// TIA Portal project "g" (V14)

(* hardware
DEVICE "S7-1200 station_1"  S7-1200 Station
   slot 0: "Rack_0"  S7-1200 Rack  Rack  V1.0
   slot 1: "PLC_1_test_mb_og_utv"  CPU 1217C DC/DC/DC  6ES7 217-1AG40-0XB0  V4.2
   slot 2: "DI 16x24VDC_1"  6ES7 221-1BH32-0XB0  V2.0
   slot 3: "CB 1241 (RS485)"  CB 1241 (RS485)  6ES7 241-1CH30-1XB0  V1.0
DEVICE "S7-1200 station_6"  S7-1200 Station
   slot 0: "Rack_0"  S7-1200 Rack  Rack  V1.0
   slot 1: "slib"  CPU 1211C DC/DC/DC  6ES7 211-1AE40-0XB0  V4.2
   slot 3: "CB 1241 (RS485)"  CB 1241 (RS485)  6ES7 241-1CH30-1XB0  V1.0
DEVICE "HMI"  TP900 Comfort
   slot 0: "TP900 Comfort"  TP900 Comfort  6AV2 124-0JC01-0AX0  14.0.1.0
   slot 1: "HMI_RT_2"  TP900 Comfort  6AV2 124-0JC01-0AX0  14.0.1.0
   slot 5: "HMI_2.IE_CP_1"  PROFINET Interface  14.0.1.0
      slot 1: "PROFINET Interface_1"  PROFINET Interface
         slot 1: "Port_1"  Port
         slot 2: "Port_2"  Port
   slot 7: "HMI_2.MPI/DP_CP_1"  MPI/DP Interface  14.0.1.0
DEVICE "S7-1200 station_2"  S7-1200 Station
   slot 0: "Rack_0"  S7-1200 Rack  Rack  V1.0
   slot 1: "PLC_1"  CPU 1211C DC/DC/DC  6ES7 211-1AE40-0XB0  V4.2
   slot 3: "CB 1241 (RS485)"  CB 1241 (RS485)  6ES7 241-1CH30-1XB0  V1.0
*)

// ===== PLC "PLC_1_test_mb_og_utv"  CPU 1217C DC/DC/DC =====

VAR_GLOBAL   // PLC tag table "Default tag table"
   "my_special_tag_name" AT %IW0 : Int;
   "tt" AT %I0.0 : Bool;
END_VAR

TYPE "mb_station_block_udt"
   STRUCT
      conf : Struct   // Configuration
         disable : Bool;   // Skip all queries
         read_only : Bool;   // Skip all write queries. (fc 5,6,15,16)
         max_comm_error : USInt := 2;   // Repeating erros before communication_error flag is set
         exec_x_quries : USInt := 1;   // Number of queries to be exec. at each loop.
      END_STRUCT;
      out : Struct   // Outputs
         error : Bool;   // All errors, including communication errors
         error_comm : Bool;   // only communication errors
         finnish : Bool;   // qid is handed over to next device.
      END_STRUCT;
      log : Struct   // Logging for development and debugging.
         connected_time : DTL;   // The time the device was connected to the bus
         disconnected_time : DTL;   // The time, if a device was disconnected to the bus
         done_cnt : UDInt;   // Successfully queries counter for this device
         error_comm_cnt : UDInt;   // Communication erros cnt.
         error_exception_cnt : UDInt;   // Failed queries counter for this device
         error_status : Word;   // Status code from mb_master or mb_client
         error_data_addr : UDInt;   // d_addr for last failed querie; handy for troubleshooting
      END_STRUCT;
      z : Struct   // Internal states.
         header_qid : UInt;   // qid value at device header
         comm_err_cnt : USInt;   // Repeating communication errors
         exec_cnt : USInt;   // Numb. of exec. q. this loop
         offset_qid : UInt := 1;   // Device query id.
         err_hold : Bool;   // Help var for .out.error
      END_STRUCT;
   END_STRUCT;
END_TYPE

// folder: mb_test

DATA_BLOCK "test_mb_t1_DB"   // DB1
{ S7_Optimized_Access := 'TRUE' }
VERSION : 0.1
// stored: InstanceOfName test_mb_1
"test_mb_1"
BEGIN
END_DATA_BLOCK

// folder: (top level)

FUNCTION_BLOCK "_read little"   // FB1, SCL
{ S7_Optimized_Access := 'TRUE' }
VERSION : 0.1
   VAR_INPUT
      mb_addr : USInt;
   END_VAR
   VAR_IN_OUT
      mb_query : "mb_query";
   END_VAR
   VAR
      sb : "mb_station_block_udt";
      data1 : Real;
      data2 : Real;
      data3 : Real;
      dommy : Bool;
      err : Int;
      pos : DInt;
   END_VAR
BEGIN

   #mb_query(mb_addr := 123,
             mode := #mb_query.c.read.holding_reg,
             data_addr := 12345,
             data_ptr := #dommy);

   IF #mb_query.Done THEN

       // #pos := "mb_pos"(mb_query := #mb_query, addr := 12345);
       #pos := UDINT_TO_DINT(12354 - #mb_query.data_addr) * 2;

       #err := READ_LITTLE(src_array := #mb_query.z.buffer,
                           dest_Variable => #data1,
                           pos := #pos);
       #err := READ_LITTLE(src_array := #mb_query.z.buffer,
                           dest_Variable => #data2,
                           pos := #pos);
       #err := READ_LITTLE(src_array := #mb_query.z.buffer,
                           dest_Variable => #data3,
                           pos := #pos);
   END_IF;
END_FUNCTION_BLOCK

FUNCTION_BLOCK "ABcounterEncoder"   // FB2, SCL
{ S7_Optimized_Access := 'TRUE' }
VERSION : 0.1
   VAR_INPUT
      pulsA : Bool;
      pulsB : Bool;
      reverce : Bool;
      factor : Real := 1.0;
   END_VAR
   VAR_OUTPUT
      pos : Real;
      uncertainPos : Bool;
   END_VAR
   VAR
      old : Struct
         pulsA : Bool;
         pulsB : Bool;
      END_STRUCT;
      cnt : DInt;
      firstScan : Bool := true;
   END_VAR
BEGIN
   // Position encoder based on two pulses which are 90 degree
   // phase shifted. 

   // TIP: Use a HSC (High speed conter) instead of this function
   // block. Using a hardware HSC will use less CPU resources.

   IF #firstScan THEN
       #uncertainPos := true;
   END_IF;

   IF #pulsA <> #old.pulsA OR #pulsB <> #old.pulsB THEN
       #cnt += SEL(G := #reverce XOR (
                    #pulsA <> NOT #old.pulsA
                    OR #pulsB <> NOT #old.pulsB),
                    IN0 := -1, IN1 := 1);
   END_IF;

   #pos := DINT_TO_REAL(#cnt) * #factor;
   #old.pulsA := #pulsA; 
   #old.pulsB := #pulsB; 
   #firstScan := false;
END_FUNCTION_BLOCK

FUNCTION_BLOCK "ABcounterCorrection"   // FB4, SCL
{ S7_Optimized_Access := 'TRUE' }
VERSION : 0.1
   VAR_INPUT
      switch : Bool;
      cnt : DInt;
   END_VAR
   VAR_OUTPUT
      deviation : DInt;
   END_VAR
   VAR_IN_OUT
      AB : "ABcounterEncoder";
   END_VAR
   VAR
      rtrig : R_TRIG;
   END_VAR
BEGIN
   #rtrig(CLK := #switch);

   // Log the max deviation
   IF NOT #AB.uncertainPos THEN
       #deviation := MAX(IN1 := #deviation, IN2 := ABS(#AB.cnt - #cnt));
   END_IF;

   IF #rtrig.Q THEN
       #AB.cnt := #cnt;
       #AB.uncertainPos := false;
   END_IF;
END_FUNCTION_BLOCK

FUNCTION "mb_get" : Void   // FC6, SCL
{ S7_Optimized_Access := 'TRUE' }
VERSION : 0.1
   VAR_INPUT
      addr : UDInt;
   END_VAR
   VAR_IN_OUT
      data_ptr : Variant;
      mb_query : "mb_query";
   END_VAR
   VAR_TEMP
      pos : DInt;
      err : Int;
   END_VAR
BEGIN
   IF #mb_query.z.run.qid_cnt = #mb_query.z.run.qid
       AND  #mb_query.Done
   THEN
       #pos := UDINT_TO_USINT(#addr - #mb_query.data_addr) * 2;
       #err := Deserialize(SRC_ARRAY := #mb_query.z.buffer,
                           DEST_VARIABLE => #data_ptr,
                           POS := #pos);
   END_IF;
END_FUNCTION

FUNCTION "mb_read_little_endian" : Void   // FC8, SCL
{ S7_Optimized_Access := 'TRUE' }
VERSION : 0.1
   VAR_INPUT
      addr : UDInt;
      n : USInt;
   END_VAR
   VAR_IN_OUT
      mb_query : "mb_query";
   END_VAR
   VAR_TEMP
      bo : Int;
      tmp : Byte;
      c : Int;
   END_VAR
BEGIN
   (* Read little endian:

      The function should be placed before a read query, and may be used 
      muliple times.

      "mb_read_little_endian"(addr := 100, n := 1, mb_query := #mb_query);
      "mb_read_little_endian"(addr := 200, n := 3, mb_query := #mb_query);

      #mb_query(mb_addr := ___MB_ADDR___,
                mode := #mb_query.c.read.holding_reg,
                data_addr := ___DATA_ADDR___,
                data_ptr := ___DATA___ );
   *) 

   IF #mb_query.z.run.qid_cnt + 1 = #mb_query.z.run.qid
       AND #mb_query.stat.done
       AND NOT #mb_query.z.run.insert
       AND NOT #mb_query.z.run.write // Read query
       AND #mb_query.conf.buffer_handler
   THEN
       #bo := UDINT_TO_INT(#addr - #mb_query.z.q.data_addr) * 2;

       FOR #c := #bo TO #bo + #n * 4 BY 4 DO
           #tmp := #mb_query.z.buffer[#bo + 0];
           #mb_query.z.buffer[#bo + 0] := #mb_query.z.buffer[#bo + 3];
           #mb_query.z.buffer[#bo + 3] := #tmp;

           #tmp := #mb_query.z.buffer[#bo + 1];
           #mb_query.z.buffer[#bo + 1] := #mb_query.z.buffer[#bo + 2];
           #mb_query.z.buffer[#bo + 2] := #tmp;
       END_FOR;
   END_IF;
END_FUNCTION

FUNCTION "mb_extra" : Bool   // FC9, SCL
{ S7_Optimized_Access := 'TRUE' }
VERSION : 0.1
   VAR_IN_OUT
      sb : "mb_station_block_udt";
      mb_query : "mb_query";
   END_VAR
BEGIN
   (* Example

   "mb_station_block_footer"(sb := #sb, mb_query := #mb_query);

   IF "mb_extra"(sb := #sb, mb_query := #mb_query) THEN
       #mb_query(mode := #mb_query.c.write.holding_reg,
                 data_addr := 12345,
                 data_ptr := ___CONFIG_PARAM___);
   END_IF;
   *)

   #mb_extra :=
   #mb_query.z.sb.sid = #mb_query.z.sb.sid_cnt
   AND NOT #sb.out.error_comm;
   // AND NOT #mb_query.stat.busy;
END_FUNCTION

ORGANIZATION_BLOCK "Main"   // OB1, SCL, ProgramCycle
TITLE = "Main Program Sweep (Cycle)"
{ S7_Optimized_Access := 'TRUE' }
VERSION : 0.1
   VAR_INPUT
      Initial_Call : Bool;   // Initial call of this OB
      Remanence : Bool;   // =True, if remanent data are available
   END_VAR
BEGIN
END_ORGANIZATION_BLOCK

// folder: mb_test

FUNCTION_BLOCK "test_mb_master"   // FB13, SCL
{ S7_Optimized_Access := 'TRUE' }
VERSION : 0.1
   VAR_INPUT
      REQ : Bool;
      MB_ADDR : UInt;
      MODE : USInt;
      DATA_ADDR : UDInt;
      DATA_LEN : UInt;
   END_VAR
   VAR_OUTPUT
      BUSY : Bool;
      ERROR : Bool;
      DONE : Bool;
      STATUS : Word;
   END_VAR
   VAR_IN_OUT
      DATA_PTR : "mb_internal_b";
   END_VAR
   VAR
      test : "test_mb_common";
   END_VAR
BEGIN
   #test(REQ := #REQ,
         MB_ADDR := #MB_ADDR,
         MODE := #MODE,
         DATA_ADDR := #DATA_ADDR,
         DATA_LEN := #DATA_LEN,
         BUSY => #BUSY,
         ERROR => #ERROR,
         DONE => #DONE,
         STATUS => #STATUS);
END_FUNCTION_BLOCK

FUNCTION_BLOCK "test_mb_common"   // FB14, SCL
{ S7_Optimized_Access := 'TRUE' }
VERSION : 0.1
   VAR_INPUT
      REQ : Bool;
      MB_ADDR : UInt;
      MODE : USInt;
      DATA_ADDR : UDInt;
      DATA_LEN : UInt;
   END_VAR
   VAR_OUTPUT
      BUSY : Bool;
      ERROR : Bool;
      DONE : Bool;
      STATUS : Word;
   END_VAR
   VAR
      fakeBus : Struct
         q : Struct
            mb_addr : UInt;
            mode : USInt;
            data_addr : UDInt;
            data_len : UInt;
         END_STRUCT;
         res : Struct
            done : Bool;
            error : Bool;
         END_STRUCT;
      END_STRUCT;
      state : Int;
      reset : Bool;
      cnt : Int;
   END_VAR
BEGIN
   // Fake query testing block

   CASE #state OF
       0:  // Wait for req.
           IF #REQ THEN
               #BUSY := true;
               #state += 1;
           END_IF;
           #cnt := 0; // Init cnt.

       1:  // Simulate some waite time
           #cnt += 1;
           #state += BOOL_TO_INT(#cnt > 5);

       2:  // Insert q-param to fake bus.
           #fakeBus.q.mb_addr := #MB_ADDR;
           #fakeBus.q.mode := #MODE;
           #fakeBus.q.data_addr := #DATA_ADDR;
           #fakeBus.q.data_len := #DATA_LEN;
           #cnt += 1; // The test device will insert resualt until next scan.

       3:  // Done or Eroor
           #fakeBus.q.mb_addr := 0;
           #fakeBus.q.mode := 0;
           #fakeBus.q.data_addr := 0;
           #fakeBus.q.data_len := 0;

           #DONE := #fakeBus.res.done;
           #ERROR := #fakeBus.res.error;
           IF NOT #DONE AND NOT #ERROR THEN
               #ERROR := true;
               #STATUS := 16#80C8;
           END_IF;
           #BUSY := false;
           #state := 0;
   END_CASE;

   IF #reset THEN
       #state := 0;
       #ERROR := false;
       #DONE := false;
       #BUSY := false;
   END_IF;

   #fakeBus.res.done := false;
   #fakeBus.res.error := false;
END_FUNCTION_BLOCK

FUNCTION_BLOCK "test_mb_client"   // FB15, SCL
{ S7_Optimized_Access := 'TRUE' }
VERSION : 0.1
   VAR_INPUT
      REQ : Bool;
      DISCONNECT : Bool;
      MB_MODE : USInt;
      DATA_ADDR : UDInt;
      DATA_LEN : UInt;
   END_VAR
   VAR_OUTPUT
      DONE : Bool;
      BUSY : Bool;
      ERROR : Bool;
      STATUS : Word;
   END_VAR
   VAR_IN_OUT
      MB_DATA_PTR : Variant;
      CONNECT : Variant;
   END_VAR
   VAR
      MB_Unit_ID : USInt;
      Connected : Bool;
      _ : Bool;
      test : "test_mb_common";
      cnt : UInt;
   END_VAR
BEGIN
   IF #DISCONNECT THEN
       #cnt := 0;
       #test.reset := true;
       #Connected := false;
   ELSE
       IF #cnt < 10 THEN
           #cnt += 1;
           #BUSY := true;
       ELSE
           #Connected := true;
           #test.reset := false;

       END_IF;
   END_IF;

   #test(REQ := #REQ,
         MB_ADDR := #MB_Unit_ID,
         MODE := #MB_MODE,
         DATA_ADDR := #DATA_ADDR,
         DATA_LEN := #DATA_LEN,
         BUSY => #BUSY,
         ERROR => #ERROR,
         DONE => #DONE,
         STATUS => #STATUS);
END_FUNCTION_BLOCK

FUNCTION_BLOCK "test_mb_1"   // FB16, SCL
{ S7_Optimized_Access := 'TRUE' }
VERSION : 0.1
   VAR_INPUT
      start : Bool;
   END_VAR
   VAR_OUTPUT
      DONE : Bool;
      ERROR : Bool;
   END_VAR
   VAR
      state : Int;
      old_state : Int;
      cnt : UInt;
      mx : UInt;
      mb_query : "mb_query";
      mb_master_1200_ctrl : "mb_master_1200_ctrl";
      mb_master_1500_ctrl : "mb_master_1200_ctrl";
      mb_client_ctrl : "mb_client_ctrl";
      mb_test_sb : Array[1..5] of "test_mb_sb1";
      mb_test_sb_fake : Array[1..5] of "test_mb_sb1_fake_device";
   END_VAR
   VAR_TEMP
      c : Int;
      dommy : Word;
   END_VAR
BEGIN
   CASE #state OF
       0:  // Wait for start signal.
           #state += BOOL_TO_INT(#start);
           #DONE := false;
           #ERROR := false;

       1:  // mb_master-1200
           #mb_test_sb[1].write1.real_1 := 0;
           #mb_test_sb[1].write1.real_2 := 0;
           #mb_test_sb[4].write1.real_1 := 0;
           #mb_test_sb[4].write1.real_2 := 0;
           #state += 1;
       2:  
           #mb_master_1200_ctrl(hardware_id := 1,
                                baud := 9600,
                                timeout := T#0s, // Auto
                                mb_query := #mb_query);

           #mb_test_sb[1].write1.real_1 := 12.34;
           #mb_test_sb[1].write1.real_2 := 56.78;
           #mb_test_sb[1]<?Sub?>(MB_ADDR := 1, mb_query := #mb_query);
           #mb_test_sb[2]<?Sub?>(MB_ADDR := 1, mb_query := #mb_query);
           #mb_test_sb[3]<?Sub?>(MB_ADDR := 1, mb_query := #mb_query);

           // Create some noice ...
           FOR #c := 0 TO UINT_TO_INT( #cnt ) MOD 7 DO
               #mb_query(mb_addr := 200, data_ptr := #dommy);
           END_FOR;

           #mb_test_sb[4].write1.real_1 := 90.12;
           #mb_test_sb[4].write1.real_2 := 34.56;
           #mb_test_sb[4]<?Sub?>(MB_ADDR := 1, mb_query := #mb_query);
           #mb_test_sb[5]<?Sub?>(MB_ADDR := 1, mb_query := #mb_query);

           FOR #c := 1 TO 5 DO
               #mb_test_sb_fake[#c]<?Sub?>(MB_ADDR := INT_TO_USINT(#c),
                                    mb_query := #mb_query,
                                    mb_test := #mb_master_1200_ctrl.master.TEST,
                                    mb_buffer := #mb_master_1200_ctrl.buffer.buffer);
           END_FOR;

           #state += BOOL_TO_INT(#cnt > 10000
                                 AND #mb_test_sb[1].read1.real_1 <> 12.34
                                 AND #mb_test_sb[1].read1.real_2 <> 56.78
                                 AND #mb_test_sb[4].read1.real_1 <> 90.12
                                 AND #mb_test_sb[4].read1.real_2 <> 34.56 );

           IF #mb_test_sb[1].read1.real_1 <> 12.34 AND #mb_test_sb[1].read1.real_1 <> 0
               OR #mb_test_sb[1].read1.real_2 <> 56.78 AND #mb_test_sb[1].read1.real_2 <> 0

               OR #mb_test_sb[4].read1.real_1 <> 90.12 AND #mb_test_sb[4].read1.real_1 <> 0
               OR #mb_test_sb[4].read1.real_2 <> 34.56 AND #mb_test_sb[4].read1.real_2 <> 0
           THEN
               #state := -1; // Error
           END_IF;

       3:  // 1500
           #mb_test_sb[3].read1.real_1 := 0;
           #state += 1;
       4:
           #mb_master_1500_ctrl(hardware_id := 1,
                                baud := 9600,
                                timeout := T#300ms,
                                mb_query := #mb_query);

           #mb_test_sb[3].write1.real_1 := 98.76;

           FOR #c := 1 TO 5 DO
               #mb_test_sb[#c]<?Sub?>(MB_ADDR := INT_TO_USINT(#c),
                               mb_query := #mb_query);
           END_FOR;

           #mb_test_sb_fake[2]<?Sub?>(MB_ADDR := INT_TO_USINT(2),
                               mb_query := #mb_query,
                               mb_test := #mb_master_1500_ctrl.master.TEST,
                               mb_buffer := #mb_master_1500_ctrl.buffer.buffer);

           #state += BOOL_TO_INT(#cnt > 10000 AND #mb_test_sb[3].read1.real_1 <> 98.76 );

           IF #mb_test_sb[3].read1.real_1 <> 98.76 AND #mb_test_sb[3].read1.real_1 <> 0 THEN
               #state := -2; // Error
               #state += 1;
           END_IF;

       5:  // Client
           #mb_test_sb[2].read1.real_1 := 0;
       6:
           #mb_client_ctrl(mb_query := #mb_query);

           #mb_test_sb[2].write1.real_1 := 0.000076;

           FOR #c := 1 TO 5 DO
               #mb_test_sb[#c]<?Sub?>(MB_ADDR := INT_TO_USINT(#c), mb_query := #mb_query);
           END_FOR;

           #mb_test_sb_fake[2]<?Sub?>(MB_ADDR := INT_TO_USINT(2),
                               mb_query := #mb_query,
                               mb_test := #mb_master_1200_ctrl.master.TEST,
                               mb_buffer := #mb_master_1200_ctrl.buffer.buffer);

           #state += BOOL_TO_INT(#cnt > 10000
                                 AND #mb_test_sb[2].read1.real_1 <> 0.000076);

           IF #mb_test_sb[2].read1.real_1 <> 0.000076 AND #mb_test_sb[2].read1.real_1 <> 0 THEN
               #state := -2; // Error
           END_IF;

       7:
           #DONE := true;
   END_CASE;

   #cnt += 1;
   IF #old_state <> #state THEN
       #cnt := 0;
   END_IF;
   #old_state := #state;

   #ERROR := #state < 0;
END_FUNCTION_BLOCK

FUNCTION_BLOCK "test_mb_comm_load"   // FB17, SCL
{ S7_Optimized_Access := 'TRUE' }
VERSION : 0.1
   VAR_INPUT
      REQ : Bool;
      PORT : Port;
      BAUD : UInt;
      PARITY : UInt;
      RESP_TO : UInt;
   END_VAR
   VAR_OUTPUT
      DONE : Bool;
      ERROR : Bool;
   END_VAR
   VAR_IN_OUT
      MB_DB : Variant;
   END_VAR
   VAR
      MB_COMM_LOAD_Instance : MB_COMM_LOAD;
      "1500" : Bool;
   END_VAR
BEGIN

   IF #"1500" THEN
       #DONE := false;
   END_IF;

   IF #REQ  
       AND #PORT <> 0 AND #BAUD <> 0 AND #PARITY <> 0 AND #RESP_TO <> 0
   THEN
       #DONE := true;
   END_IF;

   #ERROR := NOT #DONE;
END_FUNCTION_BLOCK

FUNCTION_BLOCK "test_mb_sb1_fake_device"   // FB18, SCL
{ S7_Optimized_Access := 'TRUE' }
VERSION : 0.1
   VAR_INPUT
      MB_ADDR : UInt;
   END_VAR
   VAR_IN_OUT
      mb_query : "mb_query";
      mb_test : "test_mb_common";
      mb_buffer : Array[0..250] of Byte;
   END_VAR
   VAR
      fakeBus : Struct
         q : Struct
            mb_addr : UInt;
            mode : USInt;
            data_addr : UDInt;
            data_len : UInt;
         END_STRUCT;
         res : Struct
            done : Bool;
            error : Bool;
         END_STRUCT;
      END_STRUCT;
      read1 : Struct
         real_1 : Real;
         real_2 : Real;
         udint_1 : UDInt;
      END_STRUCT;
      read2 : Struct
         x00 : Bool;
         x01 : Bool;
         x02 : Bool;
         x03 : Bool;
         x04 : Bool;
         x05 : Bool;
         x06 : Bool;
         x07 : Bool;
         x08 : Bool;
         x09 : Bool;
         x10 : Bool;
         x11 : Bool;
         x12 : Bool;
         x13 : Bool;
         x14 : Bool;
         x15 : Bool;
      END_STRUCT;
      write1 : Struct
         real_2 : Real;
         udint_1 : UDInt;
         real_1 : Real;
      END_STRUCT;
      sb : "mb_station_block_udt";
   END_VAR
   VAR_TEMP
      pos : DInt;
      "e" : Int;
   END_VAR
BEGIN
   // Simulating a device 

   IF #mb_test.fakeBus.q.mb_addr = #MB_ADDR 
       AND #mb_test.fakeBus.q.data_len > 1
   THEN
       // Read 1
       IF #mb_test.fakeBus.q.mode = #mb_query.c.read.holding_reg
           AND #mb_test.fakeBus.q.data_addr = 123
       THEN
           #"e" := Serialize(SRC_VARIABLE := #read1, DEST_ARRAY => #mb_buffer, POS := #pos);
           #mb_test.fakeBus.res.done := #"e" = 0 AND #pos / 2 = #mb_test.fakeBus.q.data_len;
       END_IF;

       // Read 2
       IF #mb_test.fakeBus.q.mode = #mb_query.c.read.holding_reg
           AND #mb_test.fakeBus.q.data_addr = 456
       THEN
           #"e" := Serialize(SRC_VARIABLE := #read2, DEST_ARRAY => #mb_buffer, POS := #pos);
           #mb_test.fakeBus.res.done := #"e" = 0 AND #pos / 2 = #mb_test.fakeBus.q.data_len;
       END_IF;

       // Write 1
       IF #mb_test.fakeBus.q.mode = #mb_query.c.write.holding_reg
           AND #mb_test.fakeBus.q.data_addr = 789
       THEN
           #"e" := Deserialize(SRC_ARRAY := #mb_buffer, DEST_VARIABLE => #write1, POS := #pos);
           #mb_test.fakeBus.res.done := #"e" = 0 AND #pos / 2 = #mb_test.fakeBus.q.data_len;
       END_IF;
   END_IF;

   #mb_test.fakeBus.res.error := NOT #mb_test.fakeBus.res.done;

   #read1.real_1 := #write1.real_1;
   #read1.real_2 := #write1.real_2;
   #read1.udint_1 := #write1.udint_1;
END_FUNCTION_BLOCK

FUNCTION_BLOCK "test_mb_sb1"   // FB19, SCL
{ S7_Optimized_Access := 'TRUE' }
VERSION : 0.1
   VAR_INPUT
      MB_ADDR : UInt;
   END_VAR
   VAR_IN_OUT
      mb_query : "mb_query";
   END_VAR
   VAR
      fakeBus : Struct
         q : Struct
            mb_addr : UInt;
            mode : USInt;
            data_addr : UDInt;
            data_len : UInt;
         END_STRUCT;
         res : Struct
            done : Bool;
            error : Bool;
         END_STRUCT;
      END_STRUCT;
      read1 : Struct
         real_1 : Real;
         real_2 : Real;
         udint_1 : UDInt;
      END_STRUCT;
      read2 : Struct
         x00 : Bool;
         x01 : Bool;
         x02 : Bool;
         x03 : Bool;
         x04 : Bool;
         x05 : Bool;
         x06 : Bool;
         x07 : Bool;
         x08 : Bool;
         x09 : Bool;
         x10 : Bool;
         x11 : Bool;
         x12 : Bool;
         x13 : Bool;
         x14 : Bool;
         x15 : Bool;
      END_STRUCT;
      write1 : Struct
         real_2 : Real;
         udint_1 : UDInt;
         real_1 : Real;
      END_STRUCT;
      sb : "mb_station_block_udt";
      q1_done_cnt : UDInt;
      q2_done_cnt : UDInt;
      q3_done_cnt : UDInt;
   END_VAR
BEGIN
   // Testing device

   "mb_station_block_header"(sb := #sb, mb_query := #mb_query);
   #mb_query.mb_addr := #MB_ADDR;

   #mb_query(mode := #mb_query.c.read.holding_reg,
             data_addr := 123,
             data_ptr := #read1);
   #q1_done_cnt += BOOL_TO_UDINT(#mb_query.Done);

   #mb_query(mode := #mb_query.c.read.holding_reg,
             data_addr := 456,
             data_ptr := #read2);
   #q2_done_cnt += BOOL_TO_UDINT(#mb_query.Done);

   #mb_query(mode := #mb_query.c.write.holding_reg,
             data_addr := 789,
             data_ptr := #write1);
   #q3_done_cnt += BOOL_TO_UDINT(#mb_query.Done);

   "mb_station_block_footer"(sb := #sb, mb_query := #mb_query);
END_FUNCTION_BLOCK

FUNCTION_BLOCK "test_mb_sb2"   // FB20, SCL
{ S7_Optimized_Access := 'TRUE' }
VERSION : 0.1
   VAR_INPUT
      MB_ADDR : UInt;
   END_VAR
   VAR_IN_OUT
      mb_query : "mb_query";
   END_VAR
   VAR
      fakeBus : Struct
         q : Struct
            mb_addr : UInt;
            mode : USInt;
            data_addr : UDInt;
            data_len : UInt;
         END_STRUCT;
         res : Struct
            done : Bool;
            error : Bool;
         END_STRUCT;
      END_STRUCT;
      read1 : Struct
         real_1 : Real;
         real_2 : Real;
         udint_1 : UDInt;
      END_STRUCT;
      read2 : Struct
         x00 : Bool;
         x01 : Bool;
         x02 : Bool;
         x03 : Bool;
         x04 : Bool;
         x05 : Bool;
         x06 : Bool;
         x07 : Bool;
         x08 : Bool;
         x09 : Bool;
         x10 : Bool;
         x11 : Bool;
         x12 : Bool;
         x13 : Bool;
         x14 : Bool;
         x15 : Bool;
      END_STRUCT;
      write1 : Struct
         real_2 : Real;
         udint_1 : UDInt;
         real_1 : Real;
      END_STRUCT;
      sb : "mb_station_block_udt";
      q1_done_cnt : UDInt;
      q2_done_cnt : UDInt;
      q3_done_cnt : UDInt;
   END_VAR
BEGIN
   // Testing device

   "mb_station_block_header"(sb := #sb, mb_query := #mb_query);
   #mb_query.mb_addr := #MB_ADDR;

   #mb_query(mode := #mb_query.c.read.holding_reg,
             data_addr := 123,
             data_ptr := #read1);
   #q1_done_cnt += BOOL_TO_UDINT(#mb_query.Done);

   #mb_query(mode := #mb_query.c.read.holding_reg,
             data_addr := 456,
             data_ptr := #read2);
   #q2_done_cnt += BOOL_TO_UDINT(#mb_query.Done);

   #mb_query(mode := #mb_query.c.write.holding_reg,
             data_addr := 789,
             data_ptr := #write1);
   #q3_done_cnt += BOOL_TO_UDINT(#mb_query.Done);

   "mb_station_block_footer"(sb := #sb, mb_query := #mb_query);
END_FUNCTION_BLOCK

FUNCTION_BLOCK "test_mb_sb2_fake_device"   // FB21, SCL
{ S7_Optimized_Access := 'TRUE' }
VERSION : 0.1
   VAR_INPUT
      MB_ADDR : UInt;
   END_VAR
   VAR_IN_OUT
      mb_query : "mb_query";
      mb_test : "test_mb_common";
      mb_buffer : Array[0..250] of Byte;
   END_VAR
   VAR
      fakeBus : Struct
         q : Struct
            mb_addr : UInt;
            mode : USInt;
            data_addr : UDInt;
            data_len : UInt;
         END_STRUCT;
         res : Struct
            done : Bool;
            error : Bool;
         END_STRUCT;
      END_STRUCT;
      read1 : Struct
         real_1 : Real;
         real_2 : Real;
         udint_1 : UDInt;
      END_STRUCT;
      read2 : Struct
         x00 : Bool;
         x01 : Bool;
         x02 : Bool;
         x03 : Bool;
         x04 : Bool;
         x05 : Bool;
         x06 : Bool;
         x07 : Bool;
         x08 : Bool;
         x09 : Bool;
         x10 : Bool;
         x11 : Bool;
         x12 : Bool;
         x13 : Bool;
         x14 : Bool;
         x15 : Bool;
      END_STRUCT;
      write1 : Struct
         real_2 : Real;
         udint_1 : UDInt;
         real_1 : Real;
      END_STRUCT;
      sb : "mb_station_block_udt";
   END_VAR
   VAR_TEMP
      pos : DInt;
      "e" : Int;
   END_VAR
BEGIN
   // Simulating a device 

   IF #mb_test.fakeBus.q.mb_addr = #MB_ADDR 
       AND #mb_test.fakeBus.q.data_len > 1
   THEN

       IF #mb_test.fakeBus.q.mode = #mb_query.c.read.input_reg
           AND #mb_test.fakeBus.q.data_addr = 123
       THEN
           #mb_test.fakeBus.res.done := false;
           #mb_test.STATUS := 16#8380; // CRC error 
       END_IF;

       IF #mb_test.fakeBus.q.mode = #mb_query.c.read.input_reg
           AND #mb_test.fakeBus.q.data_addr = 456
       THEN
           #mb_test.fakeBus.res.done := false;
           #mb_test.STATUS := 16#8384; // Data value error
       END_IF;

   END_IF;

   #mb_test.fakeBus.res.error := NOT #mb_test.fakeBus.res.done;

   #read1.real_1 := #write1.real_1;
   #read1.real_2 := #write1.real_2;
   #read1.udint_1 := #write1.udint_1;

   (* 

   Communications and configuration error messages of the instruction
   0000  No error
   80C8  Slave timeout. Check the baud rate, parity and the connectors on the slave.
   80D1  The receiver issued a flow control request to suspend an active transmission 
         and never re-enabled the transmission within the wait time.
   This  error is also generated during hardware flow control if the recipient does 
         not detect CTS within the wait time.
   80D2  The send request was aborted because no DSR signal is received from the DCE.
   80E0  The message was terminated because the receive buffer is full.
   80E1  The message was terminated as a result of a parity error.
   80E2  The message was terminated as a result of a framing error.
   80E3  The message was terminated as a result of an overrun error.
   80E4  The message was terminated as a result of the specified length exceeding the 
         total buffer size.
   8180  Invalid value for the port ID.
   8186  Invalid Modbus station address
   8188  The MODE parameter has an invalid value for a broadcast call.
   8189  Invalid data address value.
   818A  Invalid data length value.
   818B  Invalid pointer to the local data source/destination: Size not correct
   818C  The DATA_PTR parameter has an invalid pointer. Use a pointer to a bit memory 
         area or a DB with the "Standard - compatible with S7-300/400" access type.
   8200  Port is busy processing a send request


   Error messages of the Modbus protocol
   8380       CRC error 
   8381   01  Function code not supported
   8382   03  Data length error
   8383   02  Error in the data address or address outside the valid range of DATA_PTR
   8384  >03  Data value error
   8385   03  Data diagnostic code value not supported (function code 08)
   8386       Function code of the response does not match the function code of the query.
   8387       Response from wrong slave
   8388       The response of the slave to a write call is not correct. The data sent by 
              the slave does not match the query from the master.

   *)
END_FUNCTION_BLOCK

ORGANIZATION_BLOCK "test_mb_main_OB"   // OB123, SCL, ProgramCycle
TITLE = "Main Program Sweep (Cycle)"
{ S7_Optimized_Access := 'TRUE' }
VERSION : 0.1
   VAR_INPUT
      Initial_Call : Bool;   // Initial call of this OB
      Remanence : Bool;   // =True, if remanent data are available
   END_VAR
BEGIN
   "test_mb_t1_DB"();
END_ORGANIZATION_BLOCK

// ===== PLC "slib"  CPU 1211C DC/DC/DC =====

VAR_GLOBAL CONSTANT   // PLC tag table "Default tag table"
   "Handshakes.iSize" : Int := 10;
END_VAR

// ===== PLC "PLC_1"  CPU 1211C DC/DC/DC =====

// folder: Library/Alternating/Load balancer/Blocks and UDT's

TYPE "load_balancer_settings_udt"
   STRUCT
      bypass : Bool;   // Setting bypass true make all outputs enabled.
      max_devices_same_time : UInt := 65535;   // Setting, max devices that can participate at the same time
      max_diff_operating : Struct   // Max operating time between device with most and least operating time
         sec : UDInt := 4_294_967_295;
         enable : Bool;
      END_STRUCT;
      start : Struct   // Condition for starting a device
         limit : Real := 90.0;
         delay : Time := T#3M;
         force : Bool;
      END_STRUCT;
      stop : Struct   // Condition for stopping a device
         limit : Real := 20.0;
         delay : Time := T#2M;
         force : Bool;
      END_STRUCT;
      info : Struct
         input : Real;   // Block input
         total : UInt;   // Total devices
         in_operation : UInt;   // Number of devices in operation
         standby : UInt;   // Devices standby for operation
         started : UInt;   // Devices started by load balancer.
      END_STRUCT;
      boostStart : Struct   // Start correct amout of devices right away.
         enable : Bool := true;
         auto : Bool := true;   // Based on statistic on how many is usually used.
         reset : Bool;   // Reset statistics about how many devices are most frequently running.
         devices : USInt;   // Number of devices to boost start
      END_STRUCT;
   END_STRUCT;
END_TYPE

TYPE "load_balancer_device_udt"
   STRUCT
      in_operation : Bool;   // Device in operation
      available : Bool := TRUE;   // Device is available for load balancer.
      Q : Bool;   // Main output
      operation_time : UDInt;   // sec
      z : Struct   // Internal variables
         n_cnt : UDInt;   // Used for boost start. (has nothing to do with this particular device)
      END_STRUCT;
   END_STRUCT;
END_TYPE

// folder: Library/Alternating/Load balancer/Blocks and UDT's/Internal

TYPE "load_balancer_info_udt"
   STRUCT
      devices_in_operation : UInt;
      devices_standby : UInt;
      devices_started : UInt;
   END_STRUCT;
END_TYPE

// folder: Library/IO-handeling/Analog in/UDT

TYPE "alarmRealUdt"
   STRUCT
      value : Real;
      action : SInt;
      lim : Real;   // Alarm limit
      hyst : Real;   // Hysteresis
      delay : Time;   // Alarm delay
      delayEt : Time;   // delay elapsed time
      enable : Bool;   // Enable alarm
      autoAck : Bool := TRUE;   // manual acknowledge
      dobleAck : Bool;
      ack : Bool;   // acknowledge alarm
      memAck : Bool;   // Can be used for buzzer
      Q : Bool;   // output
   END_STRUCT;
END_TYPE

TYPE "analogInUdt"
   STRUCT
      filterConst : Real;   // 0=off , const for average filter.
      unitInterval : Real;   // 00.0 to 1.00 , (raw value, after running avg filter)
      sim : Bool;   // Simulate value
      forceInsideScale : Bool := true;   // Eg. in case of more then 20mA or less then 4mA.
      Error : Bool;   // Input signal out of range.
      zOldError : Bool;   // Internal variable
      ErrorTime : DTL;   // Time when the error occurred.
      errorAction : SInt := 100;   // [%]
      scaleMin : Real := 0.0;   // Scaled value for 4mA.
      scaleMax : Real := 100.0;   // Scaled value for 20mA.
      gain : Real := 1.0;   // Muliplied with the scaled value.
      offset : Real := 0.0;   // Added to "Q".
      Q : Real;   // value
   END_STRUCT;
END_TYPE

TYPE "analogInAndAlarmsUdt"
   STRUCT
      ai : "analogInUdt";
      execAiLogic : Bool := true;
      alarmL : "alarmRealUdt";
      alarmLL : "alarmRealUdt";
      alarmH : "alarmRealUdt";
      alarmHH : "alarmRealUdt";
      hmi : Struct
         copyAllSettings : Bool;
         pasteAllSettings : Bool;
         showTag : Bool;
      END_STRUCT;
   END_STRUCT;
END_TYPE

// folder: Library/IO-handeling/Analog out

TYPE "analogOutUdt"
   STRUCT
      in : Real;   // Program input
      failSafe : Bool;
      interlook : Bool;
      simEnable : Bool;
      failSafeValue : SInt := 0;   // Percent value on error, -1=keep value
      scaleMin : Real := 0.0;
      scaleMax : Real := 100.0;   // (scaleMin=0)
      simValue : Real := 0.0;
   END_STRUCT;
END_TYPE

// folder: Library/IO-handeling/Common functions

TYPE "ioGlobalUdt"
   STRUCT
      ackAllAlarms : Bool;   // Acknowledge all alarms
      disableAllSim : Bool;   // Disable all simulation of input values
      hmiShowTags : Bool;
      _ : Bool;
      totalActiveSim : UInt;   // Total active simulations
      totalActiveAlarms : UInt;   // Total active alarms
      totalUnacknowledgedAlarms : UInt;
      totalErrors : UInt;
   END_STRUCT;
END_TYPE

TYPE "alarmBoolSimpleUdt"
   STRUCT
      in : Bool;   // Input
      enable : Bool;   // Enable alarm
      autoAck : Bool := TRUE;   // Alarm will go away automaticaly when in goes false.
      dobleAck : Bool;
      ack : Bool;   // Acknowledge alarm
      memAck : Bool;   // Active alarm has been acknowledged
      Q : Bool;   // Output
   END_STRUCT;
END_TYPE

TYPE "normXAnalogUdt"
   STRUCT
      rawMin : Int := 0;
      rawMax : Int := 27648;
      errorLimMin : Int := -4864;
      errorLimMax : Int := 32512;
   END_STRUCT;
END_TYPE

// folder: Library/IO-handeling/Digital in

TYPE "digitalInUdt"
   STRUCT
      sim : Bool;   // Simulate input
      invert : Bool;   // Invert input
      Error : Bool;   // External error
      Q : Bool;   // Output
      delay : Time;   // Input delay
      delayEt : Time;
      alarm : "alarmBoolSimpleUdt";
      timeOn : DTL;
      timeOff : DTL;
   END_STRUCT;
END_TYPE

// folder: Library/IO-handeling/Digital out

TYPE "digitalOutUdt"
   STRUCT
      in : Bool;
      simEnable : Bool;
      simValue : Bool := 0;
      failSafe : Bool;
      failSafeValue : Bool;
      disableSim : Bool;
      invert : Bool;   // Invert output
   END_STRUCT;
END_TYPE

// folder: Library/Misc/operating time

TYPE "operatingTimeUdt"
   STRUCT
      operatingTime : UDInt;
      startCnt : UDInt;
      oldIn : Bool;
      oldSec : USInt;
   END_STRUCT;
END_TYPE

// folder: Library/PID

TYPE "pidUdt"
   STRUCT
      pidParam : PID_CompactControlParams;
      sp : Real;
      pv : Real;
      mv : Real;
      man : Bool;   // 0=auto
      error : Bool;
   END_STRUCT;
END_TYPE

// folder: Library/Timers/Interval

TYPE "intervalUdt"
   STRUCT
      time_between : Real;
      time_active : Real;
      time_format : SInt := 2;   // 1=ms, 2=sec, 3=min, 4=h, 5=day
      force_on : Bool;
      force_off : Bool;
      Q : Bool;
      RT : Real;
   END_STRUCT;
END_TYPE

// folder: Library/Timers/hmi timer

TYPE "timerUdt"
   STRUCT
      pt : Real;   // Preset time
      format : SInt := 2;   // 1=ms, 2=sec, 3=min, 4=h, 5=day
      RT : Real;   // Remaining time
   END_STRUCT;
END_TYPE

// folder: Library/Valves/Blocks and UDT's

TYPE "motorValveIoUdt"
   STRUCT
      in : Struct
         fullyOpen : Bool;
         fullyClosed : Bool;
         pos : Real;
         posError : Bool;
      END_STRUCT;
      out : Struct
         open : Bool;
         close : Bool;
      END_STRUCT;
      simulated : Bool;
   END_STRUCT;
END_TYPE

TYPE "motorValveConfUdt"
   STRUCT
      toggleTimeBreak : Time := T#2S;   // A short break if valve change direction.
      regModeTimeBreak : Time := T#30S;   // Wait time before a new movment when valve is regMode
      regModeMinOffset : Real := 3.0;   // Min. offset before a movment is done when valve is in regMode.
      feilSafeAction : SInt := 2;   // 0=noAction, 1=open, 2=close.
      autoReset : Bool := TRUE;   // Reset on SP change or by jog valve, else iReset need to be set true.
      simFullyOpenWithPos : Bool;   // Use the pos-signal to determined if the valve is fully open.
      simFullyClosedWithPos : Bool;   // Use the pos-signal to determined if the valve is fully closed.
      fullyOpenPosLim : Real := 98.0;   // Above this position is seen as fully open
      fullyClosedPosLim : Real := 0.7;   // Under this position is seen as fully close
      gentleOpenEnable : Bool;   // Open valve with time breaks, this may prevent damange on equipment.
      gentleCloseEnable : Bool;   // Close valve with time breaks, this may prevent damange on equipment.
      gentleAlsoOnFailSafe : Bool := TRUE;   // The gentle function will also be enabled on fail safe mode.
      gentleActivteLowLimit : Real := 15.0;   // Gentle is only activate under this limit.
      gentleTimeRun : Time := T#2S_500MS;   // Valve movment time, on gentle open or close.
      gentleTimePauseBias : Real := 4.0;   // [s] Time break between each movment on gnetle open or close.
      gentleTimePauseDelta : Real := 20.0;   // [s] The time break will increase as fracton between limit and totaly closed.
      preStop : Real := 0.3;   // Stop the movment a bit before SP is reached, so the valve will stop exactly at SP.
      endPosWithoutPreStop : Real := 3.0;   // The few last procentages on close and open, there is no preStop
      longTimeout : Time := T#4M;   // If the valve hasn't reached it's position within this time, then there is something wrong.
      quickTimeoutEnable : Bool := TRUE;   // Check at interval that the valve move towards SP.
      quickTimeoutIntervalCheaks : Time := T#8S;   // Time interval between each check.
      qucikTimeoutMinMovement : Real := 2.0;   // Min movment between each check, else error.
   END_STRUCT;
END_TYPE

TYPE "motorValveHmiUdt"
   STRUCT
      conf : "motorValveConfUdt";
      io : "motorValveIoUdt";
      error : Struct
         timeout : Bool;
         posError : Bool;
      END_STRUCT;
      cmd : Struct
         reset : Bool;
         man : Bool;   // false=>auto
         auto : Bool;
         jogOpen : Bool;
         jogClose : Bool;
         openFully : Bool;
         closeFully : Bool;
         stop : Bool;
      END_STRUCT;
      info : Struct
         regMode : Bool;   // Most be activated if valve is controlled by a PID. Makes timebreaks between each move.
         failSafe : Bool;
         interlook : Bool;
      END_STRUCT;
      SP : Real;
      operatingTime : "operatingTimeUdt";
      sim : Struct   // Simulate feedback signal
         enable : Bool;
         pos : Real;
         simByPlc : Bool;
      END_STRUCT;
      autoMan : SInt := 2;
   END_STRUCT;
END_TYPE

// folder: Library/Alternating/Load balancer

FUNCTION_BLOCK "_loadBalancer_example"   // FB14, SCL
{ S7_Optimized_Access := 'TRUE' }
VERSION : 0.1
   VAR
      load_balancer : "loadBalancer";
   END_VAR
   VAR RETAIN
      devices : Array[1..3] of "load_balancer_device_udt";
      settings : "load_balancer_settings_udt";   // Comman settings
   END_VAR
   VAR
      ___ : Bool;
      pid_output : Real;
      in_1_available : Bool;
      in_1_in_opreation : Bool;
      in_2_available : Bool;
      in_2_in_opreation : Bool;
      in_3_available : Bool;
      in_3_in_opreation : Bool;
      out_1 : Bool;
      out_2 : Bool;
      out_3 : Bool;
      out_1_value : Real;
      out_2_value : Real;
      out_3_value : Real;
   END_VAR
BEGIN
   // Load balancer example:

   // - If devices (eg. pumps) work in parallell, the function will add
   //   or remove devices to operate as the demand increase or decrease.
   // - For vfd, there should be configured a long enough ramp time to
   //   make a smooth transition when a device is added or removed for
   //   operation.
   // - More devices can be controlled, by expand the #devices array.
   // - For this theoretically example static variables bellow "___"
   //   are used, in real application the static variables would be
   //   fysical io.

   // - IMPORTANT: both #devices and #settings need to be set to retain.

   // Available: Eg. in auto, no emergensy stop, no comm.error, ready, etc.
   #devices[1].available := #in_1_available;
   #devices[2].available := #in_2_available;
   #devices[3].available := #in_3_available;

   // input:     Typically the output of a pid-controller, the "damand".
   // devices:   A array, one element for each device.
   // settings:  Can be connected to faceplate in hmi, 
   #load_balancer(input := #pid_output,
                  devices := #devices,
                  settings := #settings );
   // - Important: both #devices and #settings need to be set to retain.
   // - Open the block to see the description inside.

   // Output to devices.
   #out_1 := #devices[1].Q;
   #out_2 := #devices[2].Q;
   #out_3 := #devices[3].Q;

   // If vfd devices is controll by a vfd, then the pid_output shuld be forwared
   // to the vfd's:    
   #out_1_value := SEL(G := #devices[1].Q, IN0 := 0, IN1 := #pid_output);
   #out_2_value := SEL(G := #devices[2].Q, IN0 := 0, IN1 := #pid_output);
   #out_3_value := SEL(G := #devices[3].Q, IN0 := 0, IN1 := #pid_output);
END_FUNCTION_BLOCK

// folder: Library/Alternating/Load balancer/Blocks and UDT's

FUNCTION_BLOCK "loadBalancer"   // FB13, SCL
{ S7_Optimized_Access := 'TRUE' }
VERSION : 0.1
   VAR_INPUT
      input : Real;   // [%] Typically a output from a pid-controller.
   END_VAR
   VAR_IN_OUT
      devices : Array[*] of "load_balancer_device_udt";   // Variables for each device.
      settings : "load_balancer_settings_udt";   // Comman settings
   END_VAR
   VAR RETAIN
      conf : Struct   // Advanced configuration
         enable_operation_time_cnt : Bool := true;   // Enable operation time cnt
         at_least_one : Bool := true;   // At least one device will always be in operation
         bypass_InOperation_signal : Bool := true;   // Output control in-operation variable.
         input_zero_reset : Time := T#10M;   // All outputs will be turn off if input has been zero for this time.
         exec_boost_start_code : Bool := true;
      END_STRUCT;
   END_VAR
   VAR
      boost_start : SInt;   // Start a relative number of devices. (Negative number will stop devices)
      set : SInt := -1;   // Start a exact number of devices. (Set back to -1 right away)
      _ : Bool;
      timer_start : IEC_TIMER;
      timer_start_q : Bool;
      timer_stop : IEC_TIMER;
      timer_stop_q : Bool;
      timer_input_zero : IEC_TIMER;
      old_sec : USInt;
      ftrig_zero_input_timer : F_TRIG;
      runtime_mem1 : LReal;
      runtime_mem2 : LReal;
   END_VAR
   VAR_TEMP
      candidates : Struct
         start : Struct
            index : DInt;
            operation_time : UDInt;
         END_STRUCT;
         stop : Struct
            index : DInt;
            operation_time : UDInt;
         END_STRUCT;
      END_STRUCT;
      info : "load_balancer_info_udt";
      lower : DInt;
      upper : DInt;
      c : DInt;
      t_diff : USInt;
      oper : SInt;
      u : DInt;
      reset_timers : Bool;
      dommy : Bool;
   END_VAR
   VAR CONSTANT
      NO_CANDIDATE : DInt := 16#7fffffff;
   END_VAR
BEGIN
   (* === Load balancer ===    

   - If devices (eg. pumps) work in parallell, the function will start or stop devices
     to operate as the demand increase or decrease.
   - A devices will be added for operation, if #input is above a certain value for a
     ceratin time, eg above 90% for 50 seconds. Likewise a devices will be removed from
     operation if #input is bellow a certain value for a certain time, eg. 10% for 30
     secunds. The limits and the times are adjustable inside #settings.
   - It's the device with least operating time that will be added first, and the device
     with most operating hours will be removed from operation first.
   - #input will typically be the output of a pid-controller.
   - For vfd, there should be configured a ramp time to make a smooth transition when a
     device is added or removed for operation.
   - #devices[*].in.in_operation, is a input for fyscical feedback signal from the
     devices. this feature can be disabled by setting
     #load_balancer.conf.bypass_InOperation_signal, to true.
   - #boost_start: Make more then one devices start right away, without have to wait for
     them to start one by one. Use a negative number to stop several devies at once. One
     scan is need to start or stop each device.
   - #set: Will start or stop devies to mache number of the variable. This block will set
     the variable to -1 for the next scan.

   *)

   // If input is zero for a certain time, then all outputs is set to false.
   #timer_input_zero.TON(IN := #input = 0, PT := #conf.input_zero_reset);
   // Used to set correct number of devices from start. (Boost start)
   #ftrig_zero_input_timer(CLK := NOT #timer_input_zero.Q);

   // Default values, if the value isn't overwritten after the
   // for-loop (bellow), then there is "no candidate".
   #candidates.stop.index := #NO_CANDIDATE;
   #candidates.start.index := #NO_CANDIDATE;
   // Set to max, try find a lesser value in the for-loop bellow.
   #candidates.start.operation_time := 16#ffffffff;

   // Operating time preparing calculations:
   #runtime_mem2 += RUNTIME(#runtime_mem1);
   #t_diff := LREAL_TO_USINT(FLOOR(#runtime_mem2)); // "Overflow" if >= 1 sec.
   #runtime_mem2 -= USINT_TO_LREAL(#t_diff);

   // Boost start makes, more then one device start right away.
   IF #conf.exec_boost_start_code THEN
       "boost_start"(t_diff := #t_diff,
                     start := #ftrig_zero_input_timer.Q,
                     reset_timers => #reset_timers,
                     devices := #devices,
                     settings := #settings,
                     info := #info,
                     boost_start := #boost_start,
                     set := #set);
   END_IF;

   #lower := LOWER_BOUND(ARR := #devices, DIM := 1);
   #upper := UPPER_BOUND(ARR := #devices, DIM := 1);
   FOR #c := #lower TO #upper DO

       #devices[#c].Q := #devices[#c].Q
       (* *)AND #devices[#c].available // Disable devices that are not available. 
       (* *)AND NOT #timer_input_zero.Q // Input has not been zero for a ceratain time.
       OR #settings.bypass; // If bypass, then enable all devices.

       // If no fysical feedback signal from device for "in-operation", then
       // it's possible to bypass it.
       IF #conf.bypass_InOperation_signal THEN
           #devices[#c].in_operation := #devices[#c].Q;
       END_IF;

       REGION Candidates        
           // Candidate device to be stoped (the one that has the longest operating time)
           IF #devices[#c].Q // In use
               AND #devices[#c].operation_time >= #candidates.stop.operation_time
           THEN
               #candidates.stop.index := #c;
               #candidates.stop.operation_time := #devices[#c].operation_time;
           END_IF;

           // Candidate device to be started (the one that has the least operating time)
           IF #devices[#c].available
               AND NOT #devices[#c].Q // not allready in use
               AND #devices[#c].operation_time < #candidates.start.operation_time
           THEN
               #candidates.start.index := #c;
               #candidates.start.operation_time := #devices[#c].operation_time;
           END_IF;
       END_REGION